   1960: 'Spare_Fault_1960', class No Acknowledgement, trigger "DB302_HMI_Faults_Carrier30_Faults_2" bit 7
   1961: 'Spare_Fault_1961', class No Acknowledgement, trigger "DB302_HMI_Faults_Carrier30_Faults_2" bit 8
   1962: 'Spare_Fault_1962', class No Acknowledgement, trigger "DB302_HMI_Faults_Carrier30_Faults_2" bit 9
   1963: 'Spare_Fault_1963', class No Acknowledgement, trigger "DB302_HMI_Faults_Carrier30_Faults_2" bit 10
   1964: 'Spare_Fault_1964', class No Acknowledgement, trigger "DB302_HMI_Faults_Carrier30_Faults_2" bit 11
   1965: 'Spare_Fault_1965', class No Acknowledgement, trigger "DB302_HMI_Faults_Carrier30_Faults_2" bit 12
   1966: 'Spare_Fault_1966', class No Acknowledgement, trigger "DB302_HMI_Faults_Carrier30_Faults_2" bit 13
   1967: 'Spare_Fault_1967', class No Acknowledgement, trigger "DB302_HMI_Faults_Carrier30_Faults_2" bit 14
   1968: 'Spare_Fault_1968', class No Acknowledgement, trigger "DB302_HMI_Faults_Carrier30_Faults_2" bit 15
   1969: 'Spare_Fault_1969', class No Acknowledgement, trigger "DB302_HMI_Faults_Carrier30_Faults_3" bit 0
   1970: 'Spare_Fault_1970', class No Acknowledgement, trigger "DB302_HMI_Faults_Carrier30_Faults_3" bit 1
   1971: 'Spare_Fault_1971', class No Acknowledgement, trigger "DB302_HMI_Faults_Carrier30_Faults_3" bit 2
   1972: 'Spare_Fault_1972', class No Acknowledgement, trigger "DB302_HMI_Faults_Carrier30_Faults_3" bit 3
   1973: 'Spare_Fault_1973', class No Acknowledgement, trigger "DB302_HMI_Faults_Carrier30_Faults_3" bit 4
   1974: 'Spare_Fault_1974', class No Acknowledgement, trigger "DB302_HMI_Faults_Carrier30_Faults_3" bit 5
   1975: 'Spare_Fault_1975', class No Acknowledgement, trigger "DB302_HMI_Faults_Carrier30_Faults_3" bit 6
   1976: 'Spare_Fault_1976', class No Acknowledgement, trigger "DB302_HMI_Faults_Carrier30_Faults_3" bit 7
   1977: 'Spare_Fault_1977', class No Acknowledgement, trigger "DB302_HMI_Faults_Carrier30_Faults_3" bit 8
   1978: 'Spare_Fault_1978', class No Acknowledgement, trigger "DB302_HMI_Faults_Carrier30_Faults_3" bit 9
   1979: 'Spare_Fault_1979', class No Acknowledgement, trigger "DB302_HMI_Faults_Carrier30_Faults_3" bit 10
   1980: 'Spare_Fault_1980', class No Acknowledgement, trigger "DB302_HMI_Faults_Carrier30_Faults_3" bit 11
   1981: 'Spare_Fault_1981', class No Acknowledgement, trigger "DB302_HMI_Faults_Carrier30_Faults_3" bit 12
   1982: 'Spare_Fault_1982', class No Acknowledgement, trigger "DB302_HMI_Faults_Carrier30_Faults_3" bit 13
   1983: 'Spare_Fault_1983', class No Acknowledgement, trigger "DB302_HMI_Faults_Carrier30_Faults_3" bit 14
   1984: 'Spare_Fault_1984', class No Acknowledgement, trigger "DB302_HMI_Faults_Carrier30_Faults_3" bit 15
   1985: 'Carrier 31 Disconnect Open Power Fault DI11.0', class No Acknowledgement, trigger "DB302_HMI_Faults_Carrier31_Faults_0" bit 0
   1986: 'Carrier 31 Drive Profinet Comm Fault', class No Acknowledgement, trigger "DB302_HMI_Faults_Carrier31_Faults_0" bit 1
   1987: 'Carrier 31 Production Stop Not Reset', class No Acknowledgement, trigger "DB302_HMI_Faults_Carrier31_Faults_0" bit 2
   1988: 'Carrier 31 CB02122 Tripped', class No Acknowledgement, trigger "DB302_HMI_Faults_Carrier31_Faults_0" bit 3
   1989: 'Carrier 31 CB02123 Tripped', class No Acknowledgement, trigger "DB302_HMI_Faults_Carrier31_Faults_0" bit 4
   1990: 'Carrier 31 AUX1 CB Tripped', class No Acknowledgement, trigger "DB302_HMI_Faults_Carrier31_Faults_0" bit 5
   1991: 'Carrier 31 AUX2 CB Tripped', class No Acknowledgement, trigger "DB302_HMI_Faults_Carrier31_Faults_0" bit 6
   1992: 'Carrier 31 PLC Not Communicating', class No Acknowledgement, trigger "DB302_HMI_Faults_Carrier31_Faults_0" bit 7
   1993: 'Carrier 31 Safe Input Card Fault', class No Acknowledgement, trigger "DB302_HMI_Faults_Carrier31_Faults_0" bit 8
   1994: 'Carrier 31 Safe Output Card Fault', class No Acknowledgement, trigger "DB302_HMI_Faults_Carrier31_Faults_0" bit 9
   1995: 'Carrier 31 Standard Input Card Fault', class No Acknowledgement, trigger "DB302_HMI_Faults_Carrier31_Faults_0" bit 10
   1996: 'Carrier 31 Standard Output Card Fault', class No Acknowledgement, trigger "DB302_HMI_Faults_Carrier31_Faults_0" bit 11
   1997: 'Carrier 31 Encoder Position Fault', class No Acknowledgement, trigger "DB302_HMI_Faults_Carrier31_Faults_0" bit 12
   1998: 'Carrier 31 Encoder Internal Error', class No Acknowledgement, trigger "DB302_HMI_Faults_Carrier31_Faults_0" bit 13
   1999: 'Carrier 31 Encoder Comm Fault', class No Acknowledgement, trigger "DB302_HMI_Faults_Carrier31_Faults_0" bit 14
   2000: 'Carrier 31 HMI Comm Fault', class No Acknowledgement, trigger "DB302_HMI_Faults_Carrier31_Faults_0" bit 15
   2001: 'Carrier 31 Crash Detection Fault', class No Acknowledgement, trigger "DB302_HMI_Faults_Carrier31_Faults_1" bit 0
   2002: 'Carrier 31 Carrier Number Invalid', class No Acknowledgement, trigger "DB302_HMI_Faults_Carrier31_Faults_1" bit 1
   2003: 'Carrier 31 Drive: PROFINET configuration error', class No Acknowledgement, trigger "DB302_HMI_Faults_Carrier31_Faults_1" bit 2
   2004: 'Carrier 31 Drive: Error internal communications', class No Acknowledgement, trigger "DB302_HMI_Faults_Carrier31_Faults_1" bit 3
   2005: 'Carrier 31 Drive: Motor overtemperature', class No Acknowledgement, trigger "DB302_HMI_Faults_Carrier31_Faults_1" bit 4
   2006: 'Carrier 31 Drive: Motor overcurrent', class No Acknowledgement, trigger "DB302_HMI_Faults_Carrier31_Faults_1" bit 5
   2007: 'Carrier 31 Drive: Infeed or power unit not ready', class No Acknowledgement, trigger "DB302_HMI_Faults_Carrier31_Faults_1" bit 6
   2008: 'Carrier 31 Drive: Short-circuit/ground fault detected', class No Acknowledgement, trigger "DB302_HMI_Faults_Carrier31_Faults_1" bit 7
   2009: 'Carrier 31 Drive: PROFINET Setpoint timeout', class No Acknowledgement, trigger "DB302_HMI_Faults_Carrier31_Faults_1" bit 8
   2010: 'Carrier 31 Power unit: Overcurrent', class No Acknowledgement, trigger "DB302_HMI_Faults_Carrier31_Faults_1" bit 9
   2011: 'Carrier 31 Power unit: DC link voltage overvoltage', class No Acknowledgement, trigger "DB302_HMI_Faults_Carrier31_Faults_1" bit 10
   2012: 'Carrier 31 Power unit: DC link voltage undervoltage', class No Acknowledgement, trigger "DB302_HMI_Faults_Carrier31_Faults_1" bit 11
   2013: 'Carrier 31 Power unit: Line phase failure in main circuit', class No Acknowledgement, trigger "DB302_HMI_Faults_Carrier31_Faults_1" bit 12
   2014: 'Carrier 31 Power unit: Phase failure motor cable', class No Acknowledgement, trigger "DB302_HMI_Faults_Carrier31_Faults_1" bit 13
   2015: 'Carrier 31 Power unit: Ground fault', class No Acknowledgement, trigger "DB302_HMI_Faults_Carrier31_Faults_1" bit 14
   2016: 'Spare_Fault_2016', class No Acknowledgement, trigger "DB302_HMI_Faults_Carrier31_Faults_1" bit 15
   2017: 'Carrier 31 Motion Off Fault', class No Acknowledgement, trigger "DB302_HMI_Faults_Carrier31_Faults_2" bit 0
   2018: 'Carrier 31 Motion On Fault', class No Acknowledgement, trigger "DB302_HMI_Faults_Carrier31_Faults_2" bit 1
   2019: 'Carrier 31 Spacing Fault', class No Acknowledgement, trigger "DB302_HMI_Faults_Carrier31_Faults_2" bit 2
   2020: 'Carrier 31 Duplicate Carrier Number Fault', class No Acknowledgement, trigger "DB302_HMI_Faults_Carrier31_Faults_2" bit 3
   2021: 'Spare_Fault_2021', class No Acknowledgement, trigger "DB302_HMI_Faults_Carrier31_Faults_2" bit 4
   2022: 'Spare_Fault_2022', class No Acknowledgement, trigger "DB302_HMI_Faults_Carrier31_Faults_2" bit 5
   2023: 'Spare_Fault_2023', class No Acknowledgement, trigger "DB302_HMI_Faults_Carrier31_Faults_2" bit 6
   2024: 'Spare_Fault_2024', class No Acknowledgement, trigger "DB302_HMI_Faults_Carrier31_Faults_2" bit 7
   2025: 'Spare_Fault_2025', class No Acknowledgement, trigger "DB302_HMI_Faults_Carrier31_Faults_2" bit 8
   2026: 'Spare_Fault_2026', class No Acknowledgement, trigger "DB302_HMI_Faults_Carrier31_Faults_2" bit 9
   2027: 'Spare_Fault_2027', class No Acknowledgement, trigger "DB302_HMI_Faults_Carrier31_Faults_2" bit 10
   2028: 'Spare_Fault_2028', class No Acknowledgement, trigger "DB302_HMI_Faults_Carrier31_Faults_2" bit 11
   2029: 'Spare_Fault_2029', class No Acknowledgement, trigger "DB302_HMI_Faults_Carrier31_Faults_2" bit 12
   2030: 'Spare_Fault_2030', class No Acknowledgement, trigger "DB302_HMI_Faults_Carrier31_Faults_2" bit 13
   2031: 'Spare_Fault_2031', class No Acknowledgement, trigger "DB302_HMI_Faults_Carrier31_Faults_2" bit 14
   2032: 'Spare_Fault_2032', class No Acknowledgement, trigger "DB302_HMI_Faults_Carrier31_Faults_2" bit 15
   2033: 'Spare_Fault_2033', class No Acknowledgement, trigger "DB302_HMI_Faults_Carrier31_Faults_3" bit 0
   2034: 'Spare_Fault_2034', class No Acknowledgement, trigger "DB302_HMI_Faults_Carrier31_Faults_3" bit 1
   2035: 'Spare_Fault_2035', class No Acknowledgement, trigger "DB302_HMI_Faults_Carrier31_Faults_3" bit 2
   2036: 'Spare_Fault_2036', class No Acknowledgement, trigger "DB302_HMI_Faults_Carrier31_Faults_3" bit 3
   2037: 'Spare_Fault_2037', class No Acknowledgement, trigger "DB302_HMI_Faults_Carrier31_Faults_3" bit 4
   2038: 'Spare_Fault_2038', class No Acknowledgement, trigger "DB302_HMI_Faults_Carrier31_Faults_3" bit 5
   2039: 'Spare_Fault_2039', class No Acknowledgement, trigger "DB302_HMI_Faults_Carrier31_Faults_3" bit 6
   2040: 'Spare_Fault_2040', class No Acknowledgement, trigger "DB302_HMI_Faults_Carrier31_Faults_3" bit 7
   2041: 'Spare_Fault_2041', class No Acknowledgement, trigger "DB302_HMI_Faults_Carrier31_Faults_3" bit 8
   2042: 'Spare_Fault_2042', class No Acknowledgement, trigger "DB302_HMI_Faults_Carrier31_Faults_3" bit 9
   2043: 'Spare_Fault_2043', class No Acknowledgement, trigger "DB302_HMI_Faults_Carrier31_Faults_3" bit 10
   2044: 'Spare_Fault_2044', class No Acknowledgement, trigger "DB302_HMI_Faults_Carrier31_Faults_3" bit 11
   2045: 'Spare_Fault_2045', class No Acknowledgement, trigger "DB302_HMI_Faults_Carrier31_Faults_3" bit 12
   2046: 'Spare_Fault_2046', class No Acknowledgement, trigger "DB302_HMI_Faults_Carrier31_Faults_3" bit 13
   2047: 'Spare_Fault_2047', class No Acknowledgement, trigger "DB302_HMI_Faults_Carrier31_Faults_3" bit 14
   2048: 'Spare_Fault_2048', class No Acknowledgement, trigger "DB302_HMI_Faults_Carrier31_Faults_3" bit 15
   2049: 'Carrier 32 Disconnect Open Power Fault DI11.0', class No Acknowledgement, trigger "DB302_HMI_Faults_Carrier32_Faults_0" bit 0
   2050: 'Carrier 32 Drive Profinet Comm Fault', class No Acknowledgement, trigger "DB302_HMI_Faults_Carrier32_Faults_0" bit 1
   2051: 'Carrier 32 Production Stop Not Reset', class No Acknowledgement, trigger "DB302_HMI_Faults_Carrier32_Faults_0" bit 2
   2052: 'Carrier 32 CB02122 Tripped', class No Acknowledgement, trigger "DB302_HMI_Faults_Carrier32_Faults_0" bit 3
   2053: 'Carrier 32 CB02123 Tripped', class No Acknowledgement, trigger "DB302_HMI_Faults_Carrier32_Faults_0" bit 4
   2054: 'Carrier 32 AUX1 CB Tripped', class No Acknowledgement, trigger "DB302_HMI_Faults_Carrier32_Faults_0" bit 5
   2055: 'Carrier 32 AUX2 CB Tripped', class No Acknowledgement, trigger "DB302_HMI_Faults_Carrier32_Faults_0" bit 6
   2056: 'Carrier 32 PLC Not Communicating', class No Acknowledgement, trigger "DB302_HMI_Faults_Carrier32_Faults_0" bit 7
   2057: 'Carrier 32 Safe Input Card Fault', class No Acknowledgement, trigger "DB302_HMI_Faults_Carrier32_Faults_0" bit 8
   2058: 'Carrier 32 Safe Output Card Fault', class No Acknowledgement, trigger "DB302_HMI_Faults_Carrier32_Faults_0" bit 9
   2059: 'Carrier 32 Standard Input Card Fault', class No Acknowledgement, trigger "DB302_HMI_Faults_Carrier32_Faults_0" bit 10
   2060: 'Carrier 32 Standard Output Card Fault', class No Acknowledgement, trigger "DB302_HMI_Faults_Carrier32_Faults_0" bit 11
   2061: 'Carrier 32 Encoder Position Fault', class No Acknowledgement, trigger "DB302_HMI_Faults_Carrier32_Faults_0" bit 12
   2062: 'Carrier 32 Encoder Internal Error', class No Acknowledgement, trigger "DB302_HMI_Faults_Carrier32_Faults_0" bit 13
   2063: 'Carrier 32 Encoder Comm Fault', class No Acknowledgement, trigger "DB302_HMI_Faults_Carrier32_Faults_0" bit 14
   2064: 'Carrier 32 HMI Comm Fault', class No Acknowledgement, trigger "DB302_HMI_Faults_Carrier32_Faults_0" bit 15
   2065: 'Carrier 32 Crash Detection Fault', class No Acknowledgement, trigger "DB302_HMI_Faults_Carrier32_Faults_1" bit 0
   2066: 'Carrier 32 Carrier Number Invalid', class No Acknowledgement, trigger "DB302_HMI_Faults_Carrier32_Faults_1" bit 1
   2067: 'Carrier 32 Drive: PROFINET configuration error', class No Acknowledgement, trigger "DB302_HMI_Faults_Carrier32_Faults_1" bit 2
   2068: 'Carrier 32 Drive: Error internal communications', class No Acknowledgement, trigger "DB302_HMI_Faults_Carrier32_Faults_1" bit 3
   2069: 'Carrier 32 Drive: Motor overtemperature', class No Acknowledgement, trigger "DB302_HMI_Faults_Carrier32_Faults_1" bit 4
   2070: 'Carrier 32 Drive: Motor overcurrent', class No Acknowledgement, trigger "DB302_HMI_Faults_Carrier32_Faults_1" bit 5
   2071: 'Carrier 32 Drive: Infeed or power unit not ready', class No Acknowledgement, trigger "DB302_HMI_Faults_Carrier32_Faults_1" bit 6
   2072: 'Carrier 32 Drive: Short-circuit/ground fault detected', class No Acknowledgement, trigger "DB302_HMI_Faults_Carrier32_Faults_1" bit 7
   2073: 'Carrier 32 Drive: PROFINET Setpoint timeout', class No Acknowledgement, trigger "DB302_HMI_Faults_Carrier32_Faults_1" bit 8
   2074: 'Carrier 32 Power unit: Overcurrent', class No Acknowledgement, trigger "DB302_HMI_Faults_Carrier32_Faults_1" bit 9
   2075: 'Carrier 32 Power unit: DC link voltage overvoltage', class No Acknowledgement, trigger "DB302_HMI_Faults_Carrier32_Faults_1" bit 10
   2076: 'Carrier 32 Power unit: DC link voltage undervoltage', class No Acknowledgement, trigger "DB302_HMI_Faults_Carrier32_Faults_1" bit 11
   2077: 'Carrier 32 Power unit: Line phase failure in main circuit', class No Acknowledgement, trigger "DB302_HMI_Faults_Carrier32_Faults_1" bit 12
   2078: 'Carrier 32 Power unit: Phase failure motor cable', class No Acknowledgement, trigger "DB302_HMI_Faults_Carrier32_Faults_1" bit 13
   2079: 'Carrier 32 Power unit: Ground fault', class No Acknowledgement, trigger "DB302_HMI_Faults_Carrier32_Faults_1" bit 14
   2080: 'Spare_Fault_2080', class No Acknowledgement, trigger "DB302_HMI_Faults_Carrier32_Faults_1" bit 15
   2081: 'Carrier 32 Motion Off Fault', class No Acknowledgement, trigger "DB302_HMI_Faults_Carrier32_Faults_2" bit 0
   2082: 'Carrier 32 Motion On Fault', class No Acknowledgement, trigger "DB302_HMI_Faults_Carrier32_Faults_2" bit 1
   2083: 'Carrier 32 Spacing Fault', class No Acknowledgement, trigger "DB302_HMI_Faults_Carrier32_Faults_2" bit 2
   2084: 'Carrier 32 Duplicate Carrier Number Fault', class No Acknowledgement, trigger "DB302_HMI_Faults_Carrier32_Faults_2" bit 3
   2085: 'Spare_Fault_2085', class No Acknowledgement, trigger "DB302_HMI_Faults_Carrier32_Faults_2" bit 4
   2086: 'Spare_Fault_2086', class No Acknowledgement, trigger "DB302_HMI_Faults_Carrier32_Faults_2" bit 5
   2087: 'Spare_Fault_2087', class No Acknowledgement, trigger "DB302_HMI_Faults_Carrier32_Faults_2" bit 6
   2088: 'Spare_Fault_2088', class No Acknowledgement, trigger "DB302_HMI_Faults_Carrier32_Faults_2" bit 7
   2089: 'Spare_Fault_2089', class No Acknowledgement, trigger "DB302_HMI_Faults_Carrier32_Faults_2" bit 8
   2090: 'Spare_Fault_2090', class No Acknowledgement, trigger "DB302_HMI_Faults_Carrier32_Faults_2" bit 9
   2091: 'Spare_Fault_2091', class No Acknowledgement, trigger "DB302_HMI_Faults_Carrier32_Faults_2" bit 10
   2092: 'Spare_Fault_2092', class No Acknowledgement, trigger "DB302_HMI_Faults_Carrier32_Faults_2" bit 11
   2093: 'Spare_Fault_2093', class No Acknowledgement, trigger "DB302_HMI_Faults_Carrier32_Faults_2" bit 12
   2094: 'Spare_Fault_2094', class No Acknowledgement, trigger "DB302_HMI_Faults_Carrier32_Faults_2" bit 13
   2095: 'Spare_Fault_2095', class No Acknowledgement, trigger "DB302_HMI_Faults_Carrier32_Faults_2" bit 14
   2096: 'Spare_Fault_2096', class No Acknowledgement, trigger "DB302_HMI_Faults_Carrier32_Faults_2" bit 15
   2097: 'Spare_Fault_2097', class No Acknowledgement, trigger "DB302_HMI_Faults_Carrier32_Faults_3" bit 0
   2098: 'Spare_Fault_2098', class No Acknowledgement, trigger "DB302_HMI_Faults_Carrier32_Faults_3" bit 1
   2099: 'Spare_Fault_2099', class No Acknowledgement, trigger "DB302_HMI_Faults_Carrier32_Faults_3" bit 2
   2100: 'Spare_Fault_2100', class No Acknowledgement, trigger "DB302_HMI_Faults_Carrier32_Faults_3" bit 3
   2101: 'Spare_Fault_2101', class No Acknowledgement, trigger "DB302_HMI_Faults_Carrier32_Faults_3" bit 4
   2102: 'Spare_Fault_2102', class No Acknowledgement, trigger "DB302_HMI_Faults_Carrier32_Faults_3" bit 5
   2103: 'Spare_Fault_2103', class No Acknowledgement, trigger "DB302_HMI_Faults_Carrier32_Faults_3" bit 6
   2104: 'Spare_Fault_2104', class No Acknowledgement, trigger "DB302_HMI_Faults_Carrier32_Faults_3" bit 7
   2105: 'Spare_Fault_2105', class No Acknowledgement, trigger "DB302_HMI_Faults_Carrier32_Faults_3" bit 8
   2106: 'Spare_Fault_2106', class No Acknowledgement, trigger "DB302_HMI_Faults_Carrier32_Faults_3" bit 9
   2107: 'Spare_Fault_2107', class No Acknowledgement, trigger "DB302_HMI_Faults_Carrier32_Faults_3" bit 10
   2108: 'Spare_Fault_2108', class No Acknowledgement, trigger "DB302_HMI_Faults_Carrier32_Faults_3" bit 11
   2109: 'Spare_Fault_2109', class No Acknowledgement, trigger "DB302_HMI_Faults_Carrier32_Faults_3" bit 12
   2110: 'Spare_Fault_2110', class No Acknowledgement, trigger "DB302_HMI_Faults_Carrier32_Faults_3" bit 13
   2111: 'Spare_Fault_2111', class No Acknowledgement, trigger "DB302_HMI_Faults_Carrier32_Faults_3" bit 14
   2112: 'Spare_Fault_2112', class No Acknowledgement, trigger "DB302_HMI_Faults_Carrier32_Faults_3" bit 15
   2113: 'Carrier 33 Disconnect Open Power Fault DI11.0', class No Acknowledgement, trigger "DB302_HMI_Faults_Carrier33_Faults_0" bit 0
   2114: 'Carrier 33 Drive Profinet Comm Fault', class No Acknowledgement, trigger "DB302_HMI_Faults_Carrier33_Faults_0" bit 1
   2115: 'Carrier 33 Production Stop Not Reset', class No Acknowledgement, trigger "DB302_HMI_Faults_Carrier33_Faults_0" bit 2
   2116: 'Carrier 33 CB02122 Tripped', class No Acknowledgement, trigger "DB302_HMI_Faults_Carrier33_Faults_0" bit 3
   2117: 'Carrier 33 CB02123 Tripped', class No Acknowledgement, trigger "DB302_HMI_Faults_Carrier33_Faults_0" bit 4
   2118: 'Carrier 33 AUX1 CB Tripped', class No Acknowledgement, trigger "DB302_HMI_Faults_Carrier33_Faults_0" bit 5
   2119: 'Carrier 33 AUX2 CB Tripped', class No Acknowledgement, trigger "DB302_HMI_Faults_Carrier33_Faults_0" bit 6
   2120: 'Carrier 33 PLC Not Communicating', class No Acknowledgement, trigger "DB302_HMI_Faults_Carrier33_Faults_0" bit 7
   2121: 'Carrier 33 Safe Input Card Fault', class No Acknowledgement, trigger "DB302_HMI_Faults_Carrier33_Faults_0" bit 8
   2122: 'Carrier 33 Safe Output Card Fault', class No Acknowledgement, trigger "DB302_HMI_Faults_Carrier33_Faults_0" bit 9
   2123: 'Carrier 33 Standard Input Card Fault', class No Acknowledgement, trigger "DB302_HMI_Faults_Carrier33_Faults_0" bit 10
   2124: 'Carrier 33 Standard Output Card Fault', class No Acknowledgement, trigger "DB302_HMI_Faults_Carrier33_Faults_0" bit 11
   2125: 'Carrier 33 Encoder Position Fault', class No Acknowledgement, trigger "DB302_HMI_Faults_Carrier33_Faults_0" bit 12
   2126: 'Carrier 33 Encoder Internal Error', class No Acknowledgement, trigger "DB302_HMI_Faults_Carrier33_Faults_0" bit 13
   2127: 'Carrier 33 Encoder Comm Fault', class No Acknowledgement, trigger "DB302_HMI_Faults_Carrier33_Faults_0" bit 14
   2128: 'Carrier 33 HMI Comm Fault', class No Acknowledgement, trigger "DB302_HMI_Faults_Carrier33_Faults_0" bit 15
   2129: 'Carrier 33 Crash Detection Fault', class No Acknowledgement, trigger "DB302_HMI_Faults_Carrier33_Faults_1" bit 0
   2130: 'Carrier 33 Carrier Number Invalid', class No Acknowledgement, trigger "DB302_HMI_Faults_Carrier33_Faults_1" bit 1
   2131: 'Carrier 33 Drive: PROFINET configuration error', class No Acknowledgement, trigger "DB302_HMI_Faults_Carrier33_Faults_1" bit 2
   2132: 'Carrier 33 Drive: Error internal communications', class No Acknowledgement, trigger "DB302_HMI_Faults_Carrier33_Faults_1" bit 3
   2133: 'Carrier 33 Drive: Motor overtemperature', class No Acknowledgement, trigger "DB302_HMI_Faults_Carrier33_Faults_1" bit 4
   2134: 'Carrier 33 Drive: Motor overcurrent', class No Acknowledgement, trigger "DB302_HMI_Faults_Carrier33_Faults_1" bit 5
   2135: 'Carrier 33 Drive: Infeed or power unit not ready', class No Acknowledgement, trigger "DB302_HMI_Faults_Carrier33_Faults_1" bit 6
   2136: 'Carrier 33 Drive: Short-circuit/ground fault detected', class No Acknowledgement, trigger "DB302_HMI_Faults_Carrier33_Faults_1" bit 7
   2137: 'Carrier 33 Drive: PROFINET Setpoint timeout', class No Acknowledgement, trigger "DB302_HMI_Faults_Carrier33_Faults_1" bit 8
   2138: 'Carrier 33 Power unit: Overcurrent', class No Acknowledgement, trigger "DB302_HMI_Faults_Carrier33_Faults_1" bit 9
   2139: 'Carrier 33 Power unit: DC link voltage overvoltage', class No Acknowledgement, trigger "DB302_HMI_Faults_Carrier33_Faults_1" bit 10
   2140: 'Carrier 33 Power unit: DC link voltage undervoltage', class No Acknowledgement, trigger "DB302_HMI_Faults_Carrier33_Faults_1" bit 11
   2141: 'Carrier 33 Power unit: Line phase failure in main circuit', class No Acknowledgement, trigger "DB302_HMI_Faults_Carrier33_Faults_1" bit 12
   2142: 'Carrier 33 Power unit: Phase failure motor cable', class No Acknowledgement, trigger "DB302_HMI_Faults_Carrier33_Faults_1" bit 13
   2143: 'Carrier 33 Power unit: Ground fault', class No Acknowledgement, trigger "DB302_HMI_Faults_Carrier33_Faults_1" bit 14
   2144: 'Spare_Fault_2144', class No Acknowledgement, trigger "DB302_HMI_Faults_Carrier33_Faults_1" bit 15
   2145: 'Carrier 33 Motion Off Fault', class No Acknowledgement, trigger "DB302_HMI_Faults_Carrier33_Faults_2" bit 0
   2146: 'Carrier 33 Motion On Fault', class No Acknowledgement, trigger "DB302_HMI_Faults_Carrier33_Faults_2" bit 1
   2147: 'Carrier 33 Spacing Fault', class No Acknowledgement, trigger "DB302_HMI_Faults_Carrier33_Faults_2" bit 2
   2148: 'Carrier 33 Duplicate Carrier Number Fault', class No Acknowledgement, trigger "DB302_HMI_Faults_Carrier33_Faults_2" bit 3
   2149: 'Spare_Fault_2149', class No Acknowledgement, trigger "DB302_HMI_Faults_Carrier33_Faults_2" bit 4
   2150: 'Spare_Fault_2150', class No Acknowledgement, trigger "DB302_HMI_Faults_Carrier33_Faults_2" bit 5
   2151: 'Spare_Fault_2151', class No Acknowledgement, trigger "DB302_HMI_Faults_Carrier33_Faults_2" bit 6
   2152: 'Spare_Fault_2152', class No Acknowledgement, trigger "DB302_HMI_Faults_Carrier33_Faults_2" bit 7
   2153: 'Spare_Fault_2153', class No Acknowledgement, trigger "DB302_HMI_Faults_Carrier33_Faults_2" bit 8
   2154: 'Spare_Fault_2154', class No Acknowledgement, trigger "DB302_HMI_Faults_Carrier33_Faults_2" bit 9
   2155: 'Spare_Fault_2155', class No Acknowledgement, trigger "DB302_HMI_Faults_Carrier33_Faults_2" bit 10
   2156: 'Spare_Fault_2156', class No Acknowledgement, trigger "DB302_HMI_Faults_Carrier33_Faults_2" bit 11
   2157: 'Spare_Fault_2157', class No Acknowledgement, trigger "DB302_HMI_Faults_Carrier33_Faults_2" bit 12
   2158: 'Spare_Fault_2158', class No Acknowledgement, trigger "DB302_HMI_Faults_Carrier33_Faults_2" bit 13
   2159: 'Spare_Fault_2159', class No Acknowledgement, trigger "DB302_HMI_Faults_Carrier33_Faults_2" bit 14
   2160: 'Spare_Fault_2160', class No Acknowledgement, trigger "DB302_HMI_Faults_Carrier33_Faults_2" bit 15
   2161: 'Spare_Fault_2161', class No Acknowledgement, trigger "DB302_HMI_Faults_Carrier33_Faults_3" bit 0
   2162: 'Spare_Fault_2162', class No Acknowledgement, trigger "DB302_HMI_Faults_Carrier33_Faults_3" bit 1
   2163: 'Spare_Fault_2163', class No Acknowledgement, trigger "DB302_HMI_Faults_Carrier33_Faults_3" bit 2
   2164: 'Spare_Fault_2164', class No Acknowledgement, trigger "DB302_HMI_Faults_Carrier33_Faults_3" bit 3
   2165: 'Spare_Fault_2165', class No Acknowledgement, trigger "DB302_HMI_Faults_Carrier33_Faults_3" bit 4
   2166: 'Spare_Fault_2166', class No Acknowledgement, trigger "DB302_HMI_Faults_Carrier33_Faults_3" bit 5
   2167: 'Spare_Fault_2167', class No Acknowledgement, trigger "DB302_HMI_Faults_Carrier33_Faults_3" bit 6
   2168: 'Spare_Fault_2168', class No Acknowledgement, trigger "DB302_HMI_Faults_Carrier33_Faults_3" bit 7
   2169: 'Spare_Fault_2169', class No Acknowledgement, trigger "DB302_HMI_Faults_Carrier33_Faults_3" bit 8
   2170: 'Spare_Fault_2170', class No Acknowledgement, trigger "DB302_HMI_Faults_Carrier33_Faults_3" bit 9
   2171: 'Spare_Fault_2171', class No Acknowledgement, trigger "DB302_HMI_Faults_Carrier33_Faults_3" bit 10
   2172: 'Spare_Fault_2172', class No Acknowledgement, trigger "DB302_HMI_Faults_Carrier33_Faults_3" bit 11
   2173: 'Spare_Fault_2173', class No Acknowledgement, trigger "DB302_HMI_Faults_Carrier33_Faults_3" bit 12
   2174: 'Spare_Fault_2174', class No Acknowledgement, trigger "DB302_HMI_Faults_Carrier33_Faults_3" bit 13
   2175: 'Spare_Fault_2175', class No Acknowledgement, trigger "DB302_HMI_Faults_Carrier33_Faults_3" bit 14
   2176: 'Spare_Fault_2176', class No Acknowledgement, trigger "DB302_HMI_Faults_Carrier33_Faults_3" bit 15
   2177: 'Carrier 34 Disconnect Open Power Fault DI11.0', class No Acknowledgement, trigger "DB302_HMI_Faults_Carrier34_Faults_0" bit 0
   2178: 'Carrier 34 Drive Profinet Comm Fault', class No Acknowledgement, trigger "DB302_HMI_Faults_Carrier34_Faults_0" bit 1
   2179: 'Carrier 34 Production Stop Not Reset', class No Acknowledgement, trigger "DB302_HMI_Faults_Carrier34_Faults_0" bit 2
   2180: 'Carrier 34 CB02122 Tripped', class No Acknowledgement, trigger "DB302_HMI_Faults_Carrier34_Faults_0" bit 3
   2181: 'Carrier 34 CB02123 Tripped', class No Acknowledgement, trigger "DB302_HMI_Faults_Carrier34_Faults_0" bit 4
   2182: 'Carrier 34 AUX1 CB Tripped', class No Acknowledgement, trigger "DB302_HMI_Faults_Carrier34_Faults_0" bit 5
   2183: 'Carrier 34 AUX2 CB Tripped', class No Acknowledgement, trigger "DB302_HMI_Faults_Carrier34_Faults_0" bit 6
   2184: 'Carrier 34 PLC Not Communicating', class No Acknowledgement, trigger "DB302_HMI_Faults_Carrier34_Faults_0" bit 7
   2185: 'Carrier 34 Safe Input Card Fault', class No Acknowledgement, trigger "DB302_HMI_Faults_Carrier34_Faults_0" bit 8
   2186: 'Carrier 34 Safe Output Card Fault', class No Acknowledgement, trigger "DB302_HMI_Faults_Carrier34_Faults_0" bit 9
   2187: 'Carrier 34 Standard Input Card Fault', class No Acknowledgement, trigger "DB302_HMI_Faults_Carrier34_Faults_0" bit 10
   2188: 'Carrier 34 Standard Output Card Fault', class No Acknowledgement, trigger "DB302_HMI_Faults_Carrier34_Faults_0" bit 11
   2189: 'Carrier 34 Encoder Position Fault', class No Acknowledgement, trigger "DB302_HMI_Faults_Carrier34_Faults_0" bit 12
   2190: 'Carrier 34 Encoder Internal Error', class No Acknowledgement, trigger "DB302_HMI_Faults_Carrier34_Faults_0" bit 13
   2191: 'Carrier 34 Encoder Comm Fault', class No Acknowledgement, trigger "DB302_HMI_Faults_Carrier34_Faults_0" bit 14
   2192: 'Carrier 34 HMI Comm Fault', class No Acknowledgement, trigger "DB302_HMI_Faults_Carrier34_Faults_0" bit 15
   2193: 'Carrier 34 Crash Detection Fault', class No Acknowledgement, trigger "DB302_HMI_Faults_Carrier34_Faults_1" bit 0
   2194: 'Carrier 34 Carrier Number Invalid', class No Acknowledgement, trigger "DB302_HMI_Faults_Carrier34_Faults_1" bit 1
   2195: 'Carrier 34 Drive: PROFINET configuration error', class No Acknowledgement, trigger "DB302_HMI_Faults_Carrier34_Faults_1" bit 2
   2196: 'Carrier 34 Drive: Error internal communications', class No Acknowledgement, trigger "DB302_HMI_Faults_Carrier34_Faults_1" bit 3
   2197: 'Carrier 34 Drive: Motor overtemperature', class No Acknowledgement, trigger "DB302_HMI_Faults_Carrier34_Faults_1" bit 4
   2198: 'Carrier 34 Drive: Motor overcurrent', class No Acknowledgement, trigger "DB302_HMI_Faults_Carrier34_Faults_1" bit 5
   2199: 'Carrier 34 Drive: Infeed or power unit not ready', class No Acknowledgement, trigger "DB302_HMI_Faults_Carrier34_Faults_1" bit 6
   2200: 'Carrier 34 Drive: Short-circuit/ground fault detected', class No Acknowledgement, trigger "DB302_HMI_Faults_Carrier34_Faults_1" bit 7
   2201: 'Carrier 34 Drive: PROFINET Setpoint timeout', class No Acknowledgement, trigger "DB302_HMI_Faults_Carrier34_Faults_1" bit 8
   2202: 'Carrier 34 Power unit: Overcurrent', class No Acknowledgement, trigger "DB302_HMI_Faults_Carrier34_Faults_1" bit 9
   2203: 'Carrier 34 Power unit: DC link voltage overvoltage', class No Acknowledgement, trigger "DB302_HMI_Faults_Carrier34_Faults_1" bit 10
   2204: 'Carrier 34 Power unit: DC link voltage undervoltage', class No Acknowledgement, trigger "DB302_HMI_Faults_Carrier34_Faults_1" bit 11
   2205: 'Carrier 34 Power unit: Line phase failure in main circuit', class No Acknowledgement, trigger "DB302_HMI_Faults_Carrier34_Faults_1" bit 12
   2206: 'Carrier 34 Power unit: Phase failure motor cable', class No Acknowledgement, trigger "DB302_HMI_Faults_Carrier34_Faults_1" bit 13
   2207: 'Carrier 34 Power unit: Ground fault', class No Acknowledgement, trigger "DB302_HMI_Faults_Carrier34_Faults_1" bit 14
   2208: 'Spare_Fault_2208', class No Acknowledgement, trigger "DB302_HMI_Faults_Carrier34_Faults_1" bit 15
   2209: 'Carrier 34 Motion Off Fault', class No Acknowledgement, trigger "DB302_HMI_Faults_Carrier34_Faults_2" bit 0
   2210: 'Carrier 34 Motion On Fault', class No Acknowledgement, trigger "DB302_HMI_Faults_Carrier34_Faults_2" bit 1
   2211: 'Carrier 34 Spacing Fault', class No Acknowledgement, trigger "DB302_HMI_Faults_Carrier34_Faults_2" bit 2
   2212: 'Carrier 34 Duplicate Carrier Number Fault', class No Acknowledgement, trigger "DB302_HMI_Faults_Carrier34_Faults_2" bit 3
   2213: 'Spare_Fault_2213', class No Acknowledgement, trigger "DB302_HMI_Faults_Carrier34_Faults_2" bit 4
   2214: 'Spare_Fault_2214', class No Acknowledgement, trigger "DB302_HMI_Faults_Carrier34_Faults_2" bit 5
   2215: 'Spare_Fault_2215', class No Acknowledgement, trigger "DB302_HMI_Faults_Carrier34_Faults_2" bit 6
   2216: 'Spare_Fault_2216', class No Acknowledgement, trigger "DB302_HMI_Faults_Carrier34_Faults_2" bit 7
   2217: 'Spare_Fault_2217', class No Acknowledgement, trigger "DB302_HMI_Faults_Carrier34_Faults_2" bit 8
   2218: 'Spare_Fault_2218', class No Acknowledgement, trigger "DB302_HMI_Faults_Carrier34_Faults_2" bit 9
   2219: 'Spare_Fault_2219', class No Acknowledgement, trigger "DB302_HMI_Faults_Carrier34_Faults_2" bit 10
   2220: 'Spare_Fault_2220', class No Acknowledgement, trigger "DB302_HMI_Faults_Carrier34_Faults_2" bit 11
   2221: 'Spare_Fault_2221', class No Acknowledgement, trigger "DB302_HMI_Faults_Carrier34_Faults_2" bit 12
   2222: 'Spare_Fault_2222', class No Acknowledgement, trigger "DB302_HMI_Faults_Carrier34_Faults_2" bit 13
   2223: 'Spare_Fault_2223', class No Acknowledgement, trigger "DB302_HMI_Faults_Carrier34_Faults_2" bit 14
   2224: 'Spare_Fault_2224', class No Acknowledgement, trigger "DB302_HMI_Faults_Carrier34_Faults_2" bit 15
   2225: 'Spare_Fault_2225', class No Acknowledgement, trigger "DB302_HMI_Faults_Carrier34_Faults_3" bit 0
   2226: 'Spare_Fault_2226', class No Acknowledgement, trigger "DB302_HMI_Faults_Carrier34_Faults_3" bit 1
   2227: 'Spare_Fault_2227', class No Acknowledgement, trigger "DB302_HMI_Faults_Carrier34_Faults_3" bit 2
   2228: 'Spare_Fault_2228', class No Acknowledgement, trigger "DB302_HMI_Faults_Carrier34_Faults_3" bit 3
   2229: 'Spare_Fault_2229', class No Acknowledgement, trigger "DB302_HMI_Faults_Carrier34_Faults_3" bit 4
   2230: 'Spare_Fault_2230', class No Acknowledgement, trigger "DB302_HMI_Faults_Carrier34_Faults_3" bit 5
   2231: 'Spare_Fault_2231', class No Acknowledgement, trigger "DB302_HMI_Faults_Carrier34_Faults_3" bit 6
   2232: 'Spare_Fault_2232', class No Acknowledgement, trigger "DB302_HMI_Faults_Carrier34_Faults_3" bit 7
   2233: 'Spare_Fault_2233', class No Acknowledgement, trigger "DB302_HMI_Faults_Carrier34_Faults_3" bit 8
   2234: 'Spare_Fault_2234', class No Acknowledgement, trigger "DB302_HMI_Faults_Carrier34_Faults_3" bit 9
   2235: 'Spare_Fault_2235', class No Acknowledgement, trigger "DB302_HMI_Faults_Carrier34_Faults_3" bit 10
   2236: 'Spare_Fault_2236', class No Acknowledgement, trigger "DB302_HMI_Faults_Carrier34_Faults_3" bit 11
   2237: 'Spare_Fault_2237', class No Acknowledgement, trigger "DB302_HMI_Faults_Carrier34_Faults_3" bit 12
   2238: 'Spare_Fault_2238', class No Acknowledgement, trigger "DB302_HMI_Faults_Carrier34_Faults_3" bit 13
   2239: 'Spare_Fault_2239', class No Acknowledgement, trigger "DB302_HMI_Faults_Carrier34_Faults_3" bit 14
   2240: 'Spare_Fault_2240', class No Acknowledgement, trigger "DB302_HMI_Faults_Carrier34_Faults_3" bit 15
   2241: 'Carrier 35 Disconnect Open Power Fault DI11.0', class No Acknowledgement, trigger "DB302_HMI_Faults_Carrier35_Faults_0" bit 0
   2242: 'Carrier 35 Drive Profinet Comm Fault', class No Acknowledgement, trigger "DB302_HMI_Faults_Carrier35_Faults_0" bit 1
   2243: 'Carrier 35 Production Stop Not Reset', class No Acknowledgement, trigger "DB302_HMI_Faults_Carrier35_Faults_0" bit 2
   2244: 'Carrier 35 CB02122 Tripped', class No Acknowledgement, trigger "DB302_HMI_Faults_Carrier35_Faults_0" bit 3
   2245: 'Carrier 35 CB02123 Tripped', class No Acknowledgement, trigger "DB302_HMI_Faults_Carrier35_Faults_0" bit 4
   2246: 'Carrier 35 AUX1 CB Tripped', class No Acknowledgement, trigger "DB302_HMI_Faults_Carrier35_Faults_0" bit 5
   2247: 'Carrier 35 AUX2 CB Tripped', class No Acknowledgement, trigger "DB302_HMI_Faults_Carrier35_Faults_0" bit 6
   2248: 'Carrier 35 PLC Not Communicating', class No Acknowledgement, trigger "DB302_HMI_Faults_Carrier35_Faults_0" bit 7
   2249: 'Carrier 35 Safe Input Card Fault', class No Acknowledgement, trigger "DB302_HMI_Faults_Carrier35_Faults_0" bit 8
   2250: 'Carrier 35 Safe Output Card Fault', class No Acknowledgement, trigger "DB302_HMI_Faults_Carrier35_Faults_0" bit 9
   2251: 'Carrier 35 Standard Input Card Fault', class No Acknowledgement, trigger "DB302_HMI_Faults_Carrier35_Faults_0" bit 10
   2252: 'Carrier 35 Standard Output Card Fault', class No Acknowledgement, trigger "DB302_HMI_Faults_Carrier35_Faults_0" bit 11
   2253: 'Carrier 35 Encoder Position Fault', class No Acknowledgement, trigger "DB302_HMI_Faults_Carrier35_Faults_0" bit 12
   2254: 'Carrier 35 Encoder Internal Error', class No Acknowledgement, trigger "DB302_HMI_Faults_Carrier35_Faults_0" bit 13
   2255: 'Carrier 35 Encoder Comm Fault', class No Acknowledgement, trigger "DB302_HMI_Faults_Carrier35_Faults_0" bit 14
   2256: 'Carrier 35 HMI Comm Fault', class No Acknowledgement, trigger "DB302_HMI_Faults_Carrier35_Faults_0" bit 15
   2257: 'Carrier 35 Crash Detection Fault', class No Acknowledgement, trigger "DB302_HMI_Faults_Carrier35_Faults_1" bit 0
   2258: 'Carrier 35 Carrier Number Invalid', class No Acknowledgement, trigger "DB302_HMI_Faults_Carrier35_Faults_1" bit 1
   2259: 'Carrier 35 Drive: PROFINET configuration error', class No Acknowledgement, trigger "DB302_HMI_Faults_Carrier35_Faults_1" bit 2
   2260: 'Carrier 35 Drive: Error internal communications', class No Acknowledgement, trigger "DB302_HMI_Faults_Carrier35_Faults_1" bit 3
   2261: 'Carrier 35 Drive: Motor overtemperature', class No Acknowledgement, trigger "DB302_HMI_Faults_Carrier35_Faults_1" bit 4
   2262: 'Carrier 35 Drive: Motor overcurrent', class No Acknowledgement, trigger "DB302_HMI_Faults_Carrier35_Faults_1" bit 5
   2263: 'Carrier 35 Drive: Infeed or power unit not ready', class No Acknowledgement, trigger "DB302_HMI_Faults_Carrier35_Faults_1" bit 6
   2264: 'Carrier 35 Drive: Short-circuit/ground fault detected', class No Acknowledgement, trigger "DB302_HMI_Faults_Carrier35_Faults_1" bit 7
   2265: 'Carrier 35 Drive: PROFINET Setpoint timeout', class No Acknowledgement, trigger "DB302_HMI_Faults_Carrier35_Faults_1" bit 8
   2266: 'Carrier 35 Power unit: Overcurrent', class No Acknowledgement, trigger "DB302_HMI_Faults_Carrier35_Faults_1" bit 9
   2267: 'Carrier 35 Power unit: DC link voltage overvoltage', class No Acknowledgement, trigger "DB302_HMI_Faults_Carrier35_Faults_1" bit 10
   2268: 'Carrier 35 Power unit: DC link voltage undervoltage', class No Acknowledgement, trigger "DB302_HMI_Faults_Carrier35_Faults_1" bit 11
   2269: 'Carrier 35 Power unit: Line phase failure in main circuit', class No Acknowledgement, trigger "DB302_HMI_Faults_Carrier35_Faults_1" bit 12
   2270: 'Carrier 35 Power unit: Phase failure motor cable', class No Acknowledgement, trigger "DB302_HMI_Faults_Carrier35_Faults_1" bit 13
   2271: 'Carrier 35 Power unit: Ground fault', class No Acknowledgement, trigger "DB302_HMI_Faults_Carrier35_Faults_1" bit 14
   2272: 'Spare_Fault_2272', class No Acknowledgement, trigger "DB302_HMI_Faults_Carrier35_Faults_1" bit 15
   2273: 'Carrier 35 Motion Off Fault', class No Acknowledgement, trigger "DB302_HMI_Faults_Carrier35_Faults_2" bit 0
   2274: 'Carrier 35 Motion On Fault', class No Acknowledgement, trigger "DB302_HMI_Faults_Carrier35_Faults_2" bit 1
   2275: 'Carrier 35 Spacing Fault', class No Acknowledgement, trigger "DB302_HMI_Faults_Carrier35_Faults_2" bit 2
   2276: 'Carrier 35 Duplicate Carrier Number Fault', class No Acknowledgement, trigger "DB302_HMI_Faults_Carrier35_Faults_2" bit 3
   2277: 'Spare_Fault_2277', class No Acknowledgement, trigger "DB302_HMI_Faults_Carrier35_Faults_2" bit 4
   2278: 'Spare_Fault_2278', class No Acknowledgement, trigger "DB302_HMI_Faults_Carrier35_Faults_2" bit 5
   2279: 'Spare_Fault_2279', class No Acknowledgement, trigger "DB302_HMI_Faults_Carrier35_Faults_2" bit 6
   2280: 'Spare_Fault_2280', class No Acknowledgement, trigger "DB302_HMI_Faults_Carrier35_Faults_2" bit 7
   2281: 'Spare_Fault_2281', class No Acknowledgement, trigger "DB302_HMI_Faults_Carrier35_Faults_2" bit 8
   2282: 'Spare_Fault_2282', class No Acknowledgement, trigger "DB302_HMI_Faults_Carrier35_Faults_2" bit 9
   2283: 'Spare_Fault_2283', class No Acknowledgement, trigger "DB302_HMI_Faults_Carrier35_Faults_2" bit 10
   2284: 'Spare_Fault_2284', class No Acknowledgement, trigger "DB302_HMI_Faults_Carrier35_Faults_2" bit 11
   2285: 'Spare_Fault_2285', class No Acknowledgement, trigger "DB302_HMI_Faults_Carrier35_Faults_2" bit 12
   2286: 'Spare_Fault_2286', class No Acknowledgement, trigger "DB302_HMI_Faults_Carrier35_Faults_2" bit 13
   2287: 'Spare_Fault_2287', class No Acknowledgement, trigger "DB302_HMI_Faults_Carrier35_Faults_2" bit 14
   2288: 'Spare_Fault_2288', class No Acknowledgement, trigger "DB302_HMI_Faults_Carrier35_Faults_2" bit 15
   2289: 'Spare_Fault_2289', class No Acknowledgement, trigger "DB302_HMI_Faults_Carrier35_Faults_3" bit 0
   2290: 'Spare_Fault_2290', class No Acknowledgement, trigger "DB302_HMI_Faults_Carrier35_Faults_3" bit 1
   2291: 'Spare_Fault_2291', class No Acknowledgement, trigger "DB302_HMI_Faults_Carrier35_Faults_3" bit 2
   2292: 'Spare_Fault_2292', class No Acknowledgement, trigger "DB302_HMI_Faults_Carrier35_Faults_3" bit 3
   2293: 'Spare_Fault_2293', class No Acknowledgement, trigger "DB302_HMI_Faults_Carrier35_Faults_3" bit 4
   2294: 'Spare_Fault_2294', class No Acknowledgement, trigger "DB302_HMI_Faults_Carrier35_Faults_3" bit 5
   2295: 'Spare_Fault_2295', class No Acknowledgement, trigger "DB302_HMI_Faults_Carrier35_Faults_3" bit 6
   2296: 'Spare_Fault_2296', class No Acknowledgement, trigger "DB302_HMI_Faults_Carrier35_Faults_3" bit 7
   2297: 'Spare_Fault_2297', class No Acknowledgement, trigger "DB302_HMI_Faults_Carrier35_Faults_3" bit 8
   2298: 'Spare_Fault_2298', class No Acknowledgement, trigger "DB302_HMI_Faults_Carrier35_Faults_3" bit 9
   2299: 'Spare_Fault_2299', class No Acknowledgement, trigger "DB302_HMI_Faults_Carrier35_Faults_3" bit 10
   2300: 'Spare_Fault_2300', class No Acknowledgement, trigger "DB302_HMI_Faults_Carrier35_Faults_3" bit 11
   2301: 'Spare_Fault_2301', class No Acknowledgement, trigger "DB302_HMI_Faults_Carrier35_Faults_3" bit 12
   2302: 'Spare_Fault_2302', class No Acknowledgement, trigger "DB302_HMI_Faults_Carrier35_Faults_3" bit 13
   2303: 'Spare_Fault_2303', class No Acknowledgement, trigger "DB302_HMI_Faults_Carrier35_Faults_3" bit 14
   2304: 'Spare_Fault_2304', class No Acknowledgement, trigger "DB302_HMI_Faults_Carrier35_Faults_3" bit 15
   2305: 'Carrier36 Disconnect Open Power Fault DI11.0', class No Acknowledgement, trigger "DB302_HMI_Faults_Carrier36_Faults_0" bit 0
   2306: 'Carrier36 Drive Profinet Comm Fault', class No Acknowledgement, trigger "DB302_HMI_Faults_Carrier36_Faults_0" bit 1
   2307: 'Carrier36 Production Stop Not Reset', class No Acknowledgement, trigger "DB302_HMI_Faults_Carrier36_Faults_0" bit 2
   2308: 'Carrier36 CB02122 Tripped', class No Acknowledgement, trigger "DB302_HMI_Faults_Carrier36_Faults_0" bit 3
   2309: 'Carrier36 CB02123 Tripped', class No Acknowledgement, trigger "DB302_HMI_Faults_Carrier36_Faults_0" bit 4
   2310: 'Carrier36 AUX1 CB Tripped', class No Acknowledgement, trigger "DB302_HMI_Faults_Carrier36_Faults_0" bit 5
   2311: 'Carrier36 AUX2 CB Tripped', class No Acknowledgement, trigger "DB302_HMI_Faults_Carrier36_Faults_0" bit 6
   2312: 'Carrier36 PLC Not Communicating', class No Acknowledgement, trigger "DB302_HMI_Faults_Carrier36_Faults_0" bit 7
   2313: 'Carrier36 Safe Input Card Fault', class No Acknowledgement, trigger "DB302_HMI_Faults_Carrier36_Faults_0" bit 8
   2314: 'Carrier36 Safe Output Card Fault', class No Acknowledgement, trigger "DB302_HMI_Faults_Carrier36_Faults_0" bit 9
   2315: 'Carrier36 Standard Input Card Fault', class No Acknowledgement, trigger "DB302_HMI_Faults_Carrier36_Faults_0" bit 10
   2316: 'Carrier36 Standard Output Card Fault', class No Acknowledgement, trigger "DB302_HMI_Faults_Carrier36_Faults_0" bit 11
   2317: 'Carrier36 Encoder Position Fault', class No Acknowledgement, trigger "DB302_HMI_Faults_Carrier36_Faults_0" bit 12
   2318: 'Carrier36 Encoder Internal Error', class No Acknowledgement, trigger "DB302_HMI_Faults_Carrier36_Faults_0" bit 13
   2319: 'Carrier36 Encoder Comm Fault', class No Acknowledgement, trigger "DB302_HMI_Faults_Carrier36_Faults_0" bit 14
   2320: 'Carrier36 HMI Comm Fault', class No Acknowledgement, trigger "DB302_HMI_Faults_Carrier36_Faults_0" bit 15
   2321: 'Carrier36 Crash Detection Fault', class No Acknowledgement, trigger "DB302_HMI_Faults_Carrier36_Faults_1" bit 0
   2322: 'Carrier36 Carrier Number Invalid', class No Acknowledgement, trigger "DB302_HMI_Faults_Carrier36_Faults_1" bit 1
   2323: 'Carrier36 Drive: PROFINET configuration error', class No Acknowledgement, trigger "DB302_HMI_Faults_Carrier36_Faults_1" bit 2
   2324: 'Carrier36 Drive: Error internal communications', class No Acknowledgement, trigger "DB302_HMI_Faults_Carrier36_Faults_1" bit 3
   2325: 'Carrier36 Drive: Motor overtemperature', class No Acknowledgement, trigger "DB302_HMI_Faults_Carrier36_Faults_1" bit 4
   2326: 'Carrier36 Drive: Motor overcurrent', class No Acknowledgement, trigger "DB302_HMI_Faults_Carrier36_Faults_1" bit 5
   2327: 'Carrier36 Drive: Infeed or power unit not ready', class No Acknowledgement, trigger "DB302_HMI_Faults_Carrier36_Faults_1" bit 6
   2328: 'Carrier36 Drive: Short-circuit/ground fault detected', class No Acknowledgement, trigger "DB302_HMI_Faults_Carrier36_Faults_1" bit 7
   2329: 'Carrier36 Drive: PROFINET Setpoint timeout', class No Acknowledgement, trigger "DB302_HMI_Faults_Carrier36_Faults_1" bit 8
   2330: 'Carrier36 Power unit: Overcurrent', class No Acknowledgement, trigger "DB302_HMI_Faults_Carrier36_Faults_1" bit 9
   2331: 'Carrier36 Power unit: DC link voltage overvoltage', class No Acknowledgement, trigger "DB302_HMI_Faults_Carrier36_Faults_1" bit 10
   2332: 'Carrier36 Power unit: DC link voltage undervoltage', class No Acknowledgement, trigger "DB302_HMI_Faults_Carrier36_Faults_1" bit 11
   2333: 'Carrier36 Power unit: Line phase failure in main circuit', class No Acknowledgement, trigger "DB302_HMI_Faults_Carrier36_Faults_1" bit 12
   2334: 'Carrier36 Power unit: Phase failure motor cable', class No Acknowledgement, trigger "DB302_HMI_Faults_Carrier36_Faults_1" bit 13
   2335: 'Carrier36 Power unit: Ground fault', class No Acknowledgement, trigger "DB302_HMI_Faults_Carrier36_Faults_1" bit 14
   2336: 'Spare_Fault_2336', class No Acknowledgement, trigger "DB302_HMI_Faults_Carrier36_Faults_1" bit 15
   2337: 'Carrier36 Motion Off Fault', class No Acknowledgement, trigger "DB302_HMI_Faults_Carrier36_Faults_2" bit 0
   2338: 'Carrier36 Motion On Fault', class No Acknowledgement, trigger "DB302_HMI_Faults_Carrier36_Faults_2" bit 1
   2339: 'Carrier36 Spacing Fault', class No Acknowledgement, trigger "DB302_HMI_Faults_Carrier36_Faults_2" bit 2
   2340: 'Carrier36 Duplicate Carrier Number Fault', class No Acknowledgement, trigger "DB302_HMI_Faults_Carrier36_Faults_2" bit 3
   2341: 'Spare_Fault_2341', class No Acknowledgement, trigger "DB302_HMI_Faults_Carrier36_Faults_2" bit 4
   2342: 'Spare_Fault_2342', class No Acknowledgement, trigger "DB302_HMI_Faults_Carrier36_Faults_2" bit 5
   2343: 'Spare_Fault_2343', class No Acknowledgement, trigger "DB302_HMI_Faults_Carrier36_Faults_2" bit 6
   2344: 'Spare_Fault_2344', class No Acknowledgement, trigger "DB302_HMI_Faults_Carrier36_Faults_2" bit 7
   2345: 'Spare_Fault_2345', class No Acknowledgement, trigger "DB302_HMI_Faults_Carrier36_Faults_2" bit 8
   2346: 'Spare_Fault_2346', class No Acknowledgement, trigger "DB302_HMI_Faults_Carrier36_Faults_2" bit 9
   2347: 'Spare_Fault_2347', class No Acknowledgement, trigger "DB302_HMI_Faults_Carrier36_Faults_2" bit 10
   2348: 'Spare_Fault_2348', class No Acknowledgement, trigger "DB302_HMI_Faults_Carrier36_Faults_2" bit 11
   2349: 'Spare_Fault_2349', class No Acknowledgement, trigger "DB302_HMI_Faults_Carrier36_Faults_2" bit 12
   2350: 'Spare_Fault_2350', class No Acknowledgement, trigger "DB302_HMI_Faults_Carrier36_Faults_2" bit 13
   2351: 'Spare_Fault_2351', class No Acknowledgement, trigger "DB302_HMI_Faults_Carrier36_Faults_2" bit 14
   2352: 'Spare_Fault_2352', class No Acknowledgement, trigger "DB302_HMI_Faults_Carrier36_Faults_2" bit 15
   2353: 'Spare_Fault_2353', class No Acknowledgement, trigger "DB302_HMI_Faults_Carrier36_Faults_3" bit 0
   2354: 'Spare_Fault_2354', class No Acknowledgement, trigger "DB302_HMI_Faults_Carrier36_Faults_3" bit 1
   2355: 'Spare_Fault_2355', class No Acknowledgement, trigger "DB302_HMI_Faults_Carrier36_Faults_3" bit 2
   2356: 'Spare_Fault_2356', class No Acknowledgement, trigger "DB302_HMI_Faults_Carrier36_Faults_3" bit 3
   2357: 'Spare_Fault_2357', class No Acknowledgement, trigger "DB302_HMI_Faults_Carrier36_Faults_3" bit 4
   2358: 'Spare_Fault_2358', class No Acknowledgement, trigger "DB302_HMI_Faults_Carrier36_Faults_3" bit 5
   2359: 'Spare_Fault_2359', class No Acknowledgement, trigger "DB302_HMI_Faults_Carrier36_Faults_3" bit 6
   2360: 'Spare_Fault_2360', class No Acknowledgement, trigger "DB302_HMI_Faults_Carrier36_Faults_3" bit 7
   2361: 'Spare_Fault_2361', class No Acknowledgement, trigger "DB302_HMI_Faults_Carrier36_Faults_3" bit 8
   2362: 'Spare_Fault_2362', class No Acknowledgement, trigger "DB302_HMI_Faults_Carrier36_Faults_3" bit 9
   2363: 'Spare_Fault_2363', class No Acknowledgement, trigger "DB302_HMI_Faults_Carrier36_Faults_3" bit 10
   2364: 'Spare_Fault_2364', class No Acknowledgement, trigger "DB302_HMI_Faults_Carrier36_Faults_3" bit 11
   2365: 'Spare_Fault_2365', class No Acknowledgement, trigger "DB302_HMI_Faults_Carrier36_Faults_3" bit 12
   2366: 'Spare_Fault_2366', class No Acknowledgement, trigger "DB302_HMI_Faults_Carrier36_Faults_3" bit 13
   2367: 'Spare_Fault_2367', class No Acknowledgement, trigger "DB302_HMI_Faults_Carrier36_Faults_3" bit 14
   2368: 'Spare_Fault_2368', class No Acknowledgement, trigger "DB302_HMI_Faults_Carrier36_Faults_3" bit 15
   2369: 'Carrier 37 Disconnect Open Power Fault DI11.0', class No Acknowledgement, trigger "DB302_HMI_Faults_Carrier37_Faults_0" bit 0
   2370: 'Carrier 37 Drive Profinet Comm Fault', class No Acknowledgement, trigger "DB302_HMI_Faults_Carrier37_Faults_0" bit 1
   2371: 'Carrier 37 Production Stop Not Reset', class No Acknowledgement, trigger "DB302_HMI_Faults_Carrier37_Faults_0" bit 2
   2372: 'Carrier 37 CB02122 Tripped', class No Acknowledgement, trigger "DB302_HMI_Faults_Carrier37_Faults_0" bit 3
   2373: 'Carrier 37 CB02123 Tripped', class No Acknowledgement, trigger "DB302_HMI_Faults_Carrier37_Faults_0" bit 4
   2374: 'Carrier 37 AUX1 CB Tripped', class No Acknowledgement, trigger "DB302_HMI_Faults_Carrier37_Faults_0" bit 5
   2375: 'Carrier 37 AUX2 CB Tripped', class No Acknowledgement, trigger "DB302_HMI_Faults_Carrier37_Faults_0" bit 6
   2376: 'Carrier 37 PLC Not Communicating', class No Acknowledgement, trigger "DB302_HMI_Faults_Carrier37_Faults_0" bit 7
   2377: 'Carrier 37 Safe Input Card Fault', class No Acknowledgement, trigger "DB302_HMI_Faults_Carrier37_Faults_0" bit 8
   2378: 'Carrier 37 Safe Output Card Fault', class No Acknowledgement, trigger "DB302_HMI_Faults_Carrier37_Faults_0" bit 9
   2379: 'Carrier 37 Standard Input Card Fault', class No Acknowledgement, trigger "DB302_HMI_Faults_Carrier37_Faults_0" bit 10
   2380: 'Carrier 37 Standard Output Card Fault', class No Acknowledgement, trigger "DB302_HMI_Faults_Carrier37_Faults_0" bit 11
   2381: 'Carrier 37 Encoder Position Fault', class No Acknowledgement, trigger "DB302_HMI_Faults_Carrier37_Faults_0" bit 12
   2382: 'Carrier 37 Encoder Internal Error', class No Acknowledgement, trigger "DB302_HMI_Faults_Carrier37_Faults_0" bit 13
